(* Logix 5000 project; controller PLC_MCC1300_75F1 vendor 1 type 14 code 166 rev 32.11; software revision 32.04; part 49 of 83 *)
(* tags used below, declared in another part *)
   GP_ConversionXY : GP_ConversionXY;
   M30xTrimWheel : MAC_TrimmingWheels[5];
   M30xTrimWheel_HMR : MAC_TrimmingWheels_HMR[5];
   M30xTrimWheel_HMW : MAC_TrimmingWheels_HMW[5];
   M310B : MAC_Conveyor;
   M310B_ALM : MAC_Conveyor_ALM;
   M310B_Data : UDT_Convoy_SL;
   M310B_SpaceConv_Utilities : SpaceConv_Utilities;
   TMP_dIndex : DINT;
   TMP_rActualValue_cmm : REAL;
   xAlwaysON : BOOL;
   xDebugOFF : BOOL;
   Z401 : MAC_Zone;
(* MainProgram, continued *)

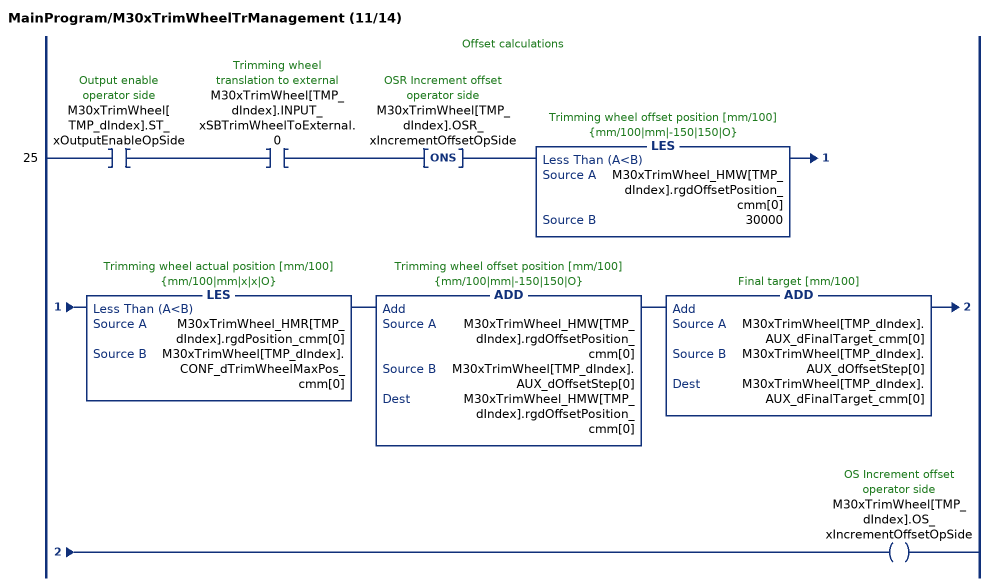
   [picture p745: MainProgram/M30xTrimWheelTrManagement rungs 25-25]
   // Offset calculations
   25: XIC(M30xTrimWheel[TMP_dIndex].ST_xOutputEnableOpSide)XIC(M30xTrimWheel[TMP_dIndex].INPUT_xSBTrimWheelToExternal.0)ONS(M30xTrimWheel[TMP_dIndex].OSR_xIncrementOffsetOpSide)LES(M30xTrimWheel_HMW[TMP_dIndex].rgdOffsetPosition_cmm[0],30000)LES(M30xTrimWheel_HMR[TMP_dIndex].rgdPosition_cmm[0],M30xTrimWheel[TMP_dIndex].CONF_dTrimWheelMaxPos_cmm[0])ADD(M30xTrimWheel_HMW[TMP_dIndex].rgdOffsetPosition_cmm[0],M30xTrimWheel[TMP_dIndex].AUX_dOffsetStep[0],M30xTrimWheel_HMW[TMP_dIndex].rgdOffsetPosition_cmm[0])ADD(M30xTrimWheel[TMP_dIndex].AUX_dFinalTarget_cmm[0],M30xTrimWheel[TMP_dIndex].AUX_dOffsetStep[0],M30xTrimWheel[TMP_dIndex].AUX_dFinalTarget_cmm[0])OTE(M30xTrimWheel[TMP_dIndex].OS_xIncrementOffsetOpSide);
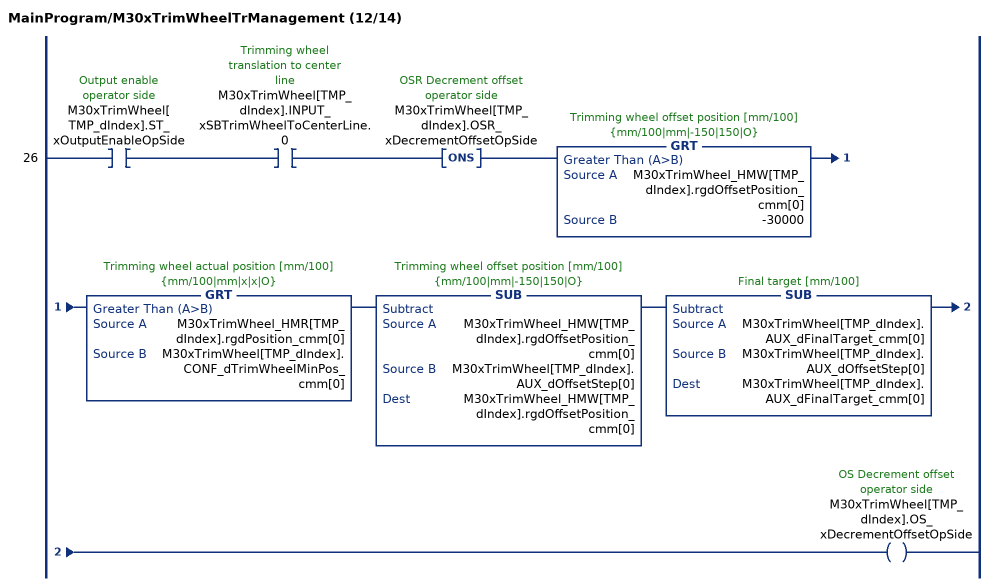
   26: XIC(M30xTrimWheel[TMP_dIndex].ST_xOutputEnableOpSide)XIC(M30xTrimWheel[TMP_dIndex].INPUT_xSBTrimWheelToCenterLine.0)ONS(M30xTrimWheel[TMP_dIndex].OSR_xDecrementOffsetOpSide)GRT(M30xTrimWheel_HMW[TMP_dIndex].rgdOffsetPosition_cmm[0],-30000)GRT(M30xTrimWheel_HMR[TMP_dIndex].rgdPosition_cmm[0],M30xTrimWheel[TMP_dIndex].CONF_dTrimWheelMinPos_cmm[0])SUB(M30xTrimWheel_HMW[TMP_dIndex].rgdOffsetPosition_cmm[0],M30xTrimWheel[TMP_dIndex].AUX_dOffsetStep[0],M30xTrimWheel_HMW[TMP_dIndex].rgdOffsetPosition_cmm[0])SUB(M30xTrimWheel[TMP_dIndex].AUX_dFinalTarget_cmm[0],M30xTrimWheel[TMP_dIndex].AUX_dOffsetStep[0],M30xTrimWheel[TMP_dIndex].AUX_dFinalTarget_cmm[0])OTE(M30xTrimWheel[TMP_dIndex].OS_xDecrementOffsetOpSide);
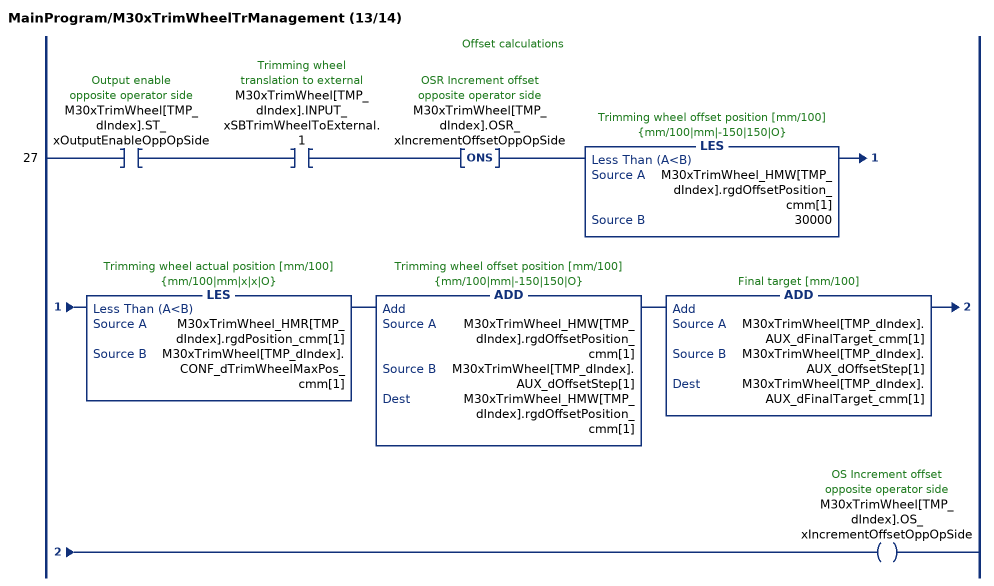
   // Offset calculations
   27: XIC(M30xTrimWheel[TMP_dIndex].ST_xOutputEnableOppOpSide)XIC(M30xTrimWheel[TMP_dIndex].INPUT_xSBTrimWheelToExternal.1)ONS(M30xTrimWheel[TMP_dIndex].OSR_xIncrementOffsetOppOpSide)LES(M30xTrimWheel_HMW[TMP_dIndex].rgdOffsetPosition_cmm[1],30000)LES(M30xTrimWheel_HMR[TMP_dIndex].rgdPosition_cmm[1],M30xTrimWheel[TMP_dIndex].CONF_dTrimWheelMaxPos_cmm[1])ADD(M30xTrimWheel_HMW[TMP_dIndex].rgdOffsetPosition_cmm[1],M30xTrimWheel[TMP_dIndex].AUX_dOffsetStep[1],M30xTrimWheel_HMW[TMP_dIndex].rgdOffsetPosition_cmm[1])ADD(M30xTrimWheel[TMP_dIndex].AUX_dFinalTarget_cmm[1],M30xTrimWheel[TMP_dIndex].AUX_dOffsetStep[1],M30xTrimWheel[TMP_dIndex].AUX_dFinalTarget_cmm[1])OTE(M30xTrimWheel[TMP_dIndex].OS_xIncrementOffsetOppOpSide);
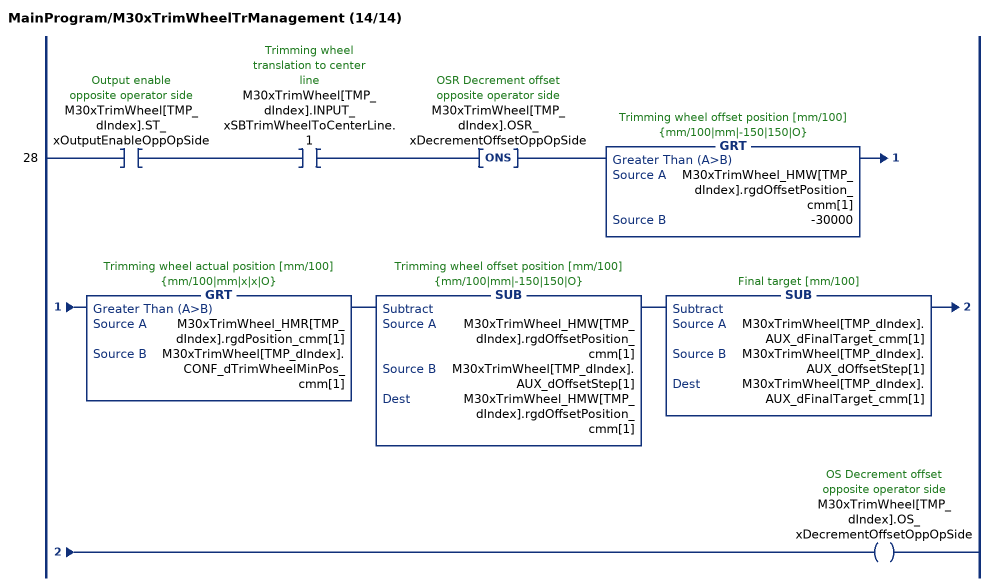
   28: XIC(M30xTrimWheel[TMP_dIndex].ST_xOutputEnableOppOpSide)XIC(M30xTrimWheel[TMP_dIndex].INPUT_xSBTrimWheelToCenterLine.1)ONS(M30xTrimWheel[TMP_dIndex].OSR_xDecrementOffsetOppOpSide)GRT(M30xTrimWheel_HMW[TMP_dIndex].rgdOffsetPosition_cmm[1],-30000)GRT(M30xTrimWheel_HMR[TMP_dIndex].rgdPosition_cmm[1],M30xTrimWheel[TMP_dIndex].CONF_dTrimWheelMinPos_cmm[1])SUB(M30xTrimWheel_HMW[TMP_dIndex].rgdOffsetPosition_cmm[1],M30xTrimWheel[TMP_dIndex].AUX_dOffsetStep[1],M30xTrimWheel_HMW[TMP_dIndex].rgdOffsetPosition_cmm[1])SUB(M30xTrimWheel[TMP_dIndex].AUX_dFinalTarget_cmm[1],M30xTrimWheel[TMP_dIndex].AUX_dOffsetStep[1],M30xTrimWheel[TMP_dIndex].AUX_dFinalTarget_cmm[1])OTE(M30xTrimWheel[TMP_dIndex].OS_xDecrementOffsetOppOpSide);
END_ROUTINE

ROUTINE M30xTrimWheelTrOppOpSide_Logic   (* ladder *)
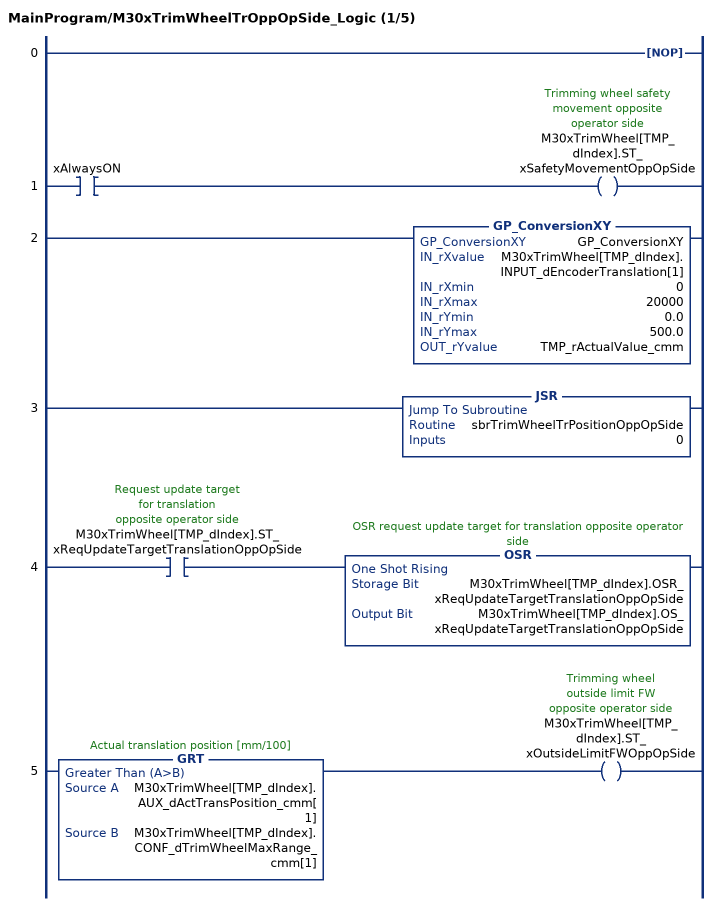
   0: NOP();
   1: XIC(xAlwaysON)OTE(M30xTrimWheel[TMP_dIndex].ST_xSafetyMovementOppOpSide);
   2: GP_ConversionXY(GP_ConversionXY,M30xTrimWheel[TMP_dIndex].INPUT_dEncoderTranslation[1],0,20000,0.0,500.0,TMP_rActualValue_cmm);
   3: JSR(sbrTrimWheelTrPositionOppOpSide,0);
   4: XIC(M30xTrimWheel[TMP_dIndex].ST_xReqUpdateTargetTranslationOppOpSide)OSR(M30xTrimWheel[TMP_dIndex].OSR_xReqUpdateTargetTranslationOppOpSide,M30xTrimWheel[TMP_dIndex].OS_xReqUpdateTargetTranslationOppOpSide);
   5: GRT(M30xTrimWheel[TMP_dIndex].AUX_dActTransPosition_cmm[1],M30xTrimWheel[TMP_dIndex].CONF_dTrimWheelMaxRange_cmm[1])OTE(M30xTrimWheel[TMP_dIndex].ST_xOutsideLimitFWOppOpSide);
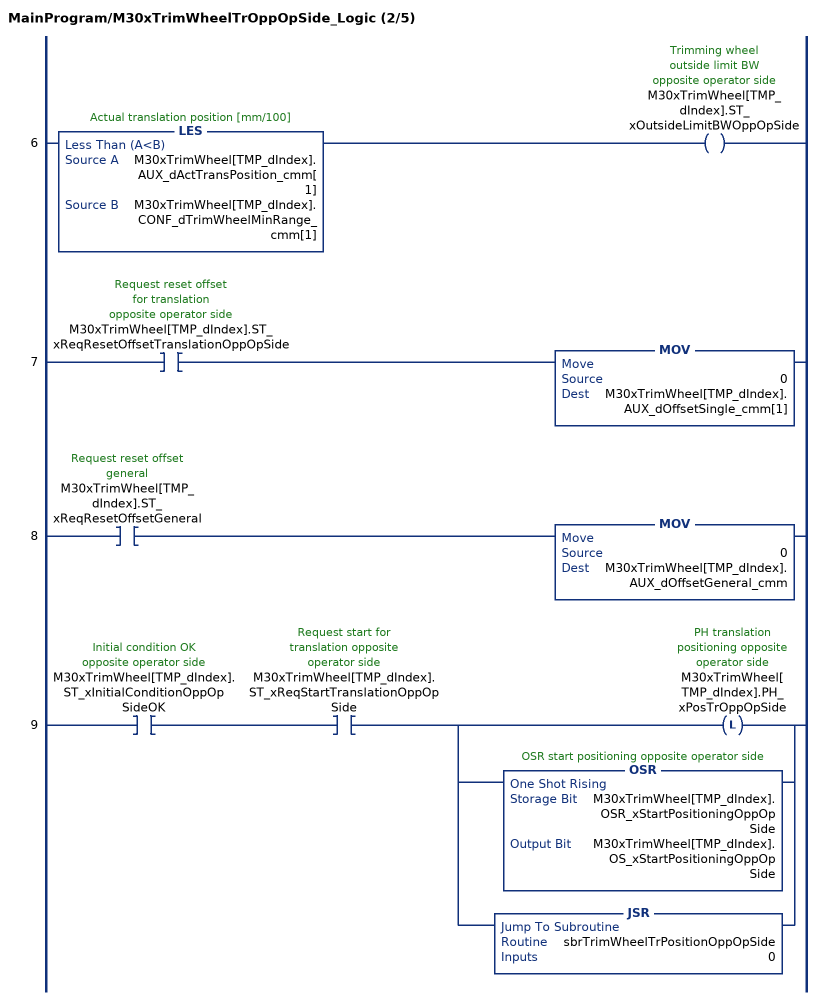
   6: LES(M30xTrimWheel[TMP_dIndex].AUX_dActTransPosition_cmm[1],M30xTrimWheel[TMP_dIndex].CONF_dTrimWheelMinRange_cmm[1])OTE(M30xTrimWheel[TMP_dIndex].ST_xOutsideLimitBWOppOpSide);
   7: XIC(M30xTrimWheel[TMP_dIndex].ST_xReqResetOffsetTranslationOppOpSide)MOV(0,M30xTrimWheel[TMP_dIndex].AUX_dOffsetSingle_cmm[1]);
   8: XIC(M30xTrimWheel[TMP_dIndex].ST_xReqResetOffsetGeneral)MOV(0,M30xTrimWheel[TMP_dIndex].AUX_dOffsetGeneral_cmm);
   9: XIC(M30xTrimWheel[TMP_dIndex].ST_xInitialConditionOppOpSideOK)XIC(M30xTrimWheel[TMP_dIndex].ST_xReqStartTranslationOppOpSide)[OTL(M30xTrimWheel[TMP_dIndex].PH_xPosTrOppOpSide) ,OSR(M30xTrimWheel[TMP_dIndex].OSR_xStartPositioningOppOpSide,M30xTrimWheel[TMP_dIndex].OS_xStartPositioningOppOpSide) ,JSR(sbrTrimWheelTrPositionOppOpSide,0) ];
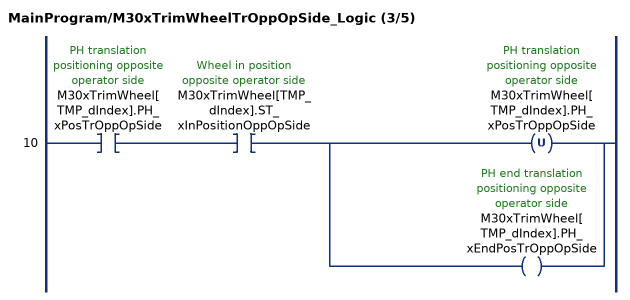
   10: XIC(M30xTrimWheel[TMP_dIndex].PH_xPosTrOppOpSide)XIC(M30xTrimWheel[TMP_dIndex].ST_xInPositionOppOpSide)[OTU(M30xTrimWheel[TMP_dIndex].PH_xPosTrOppOpSide) ,OTE(M30xTrimWheel[TMP_dIndex].PH_xEndPosTrOppOpSide) ];
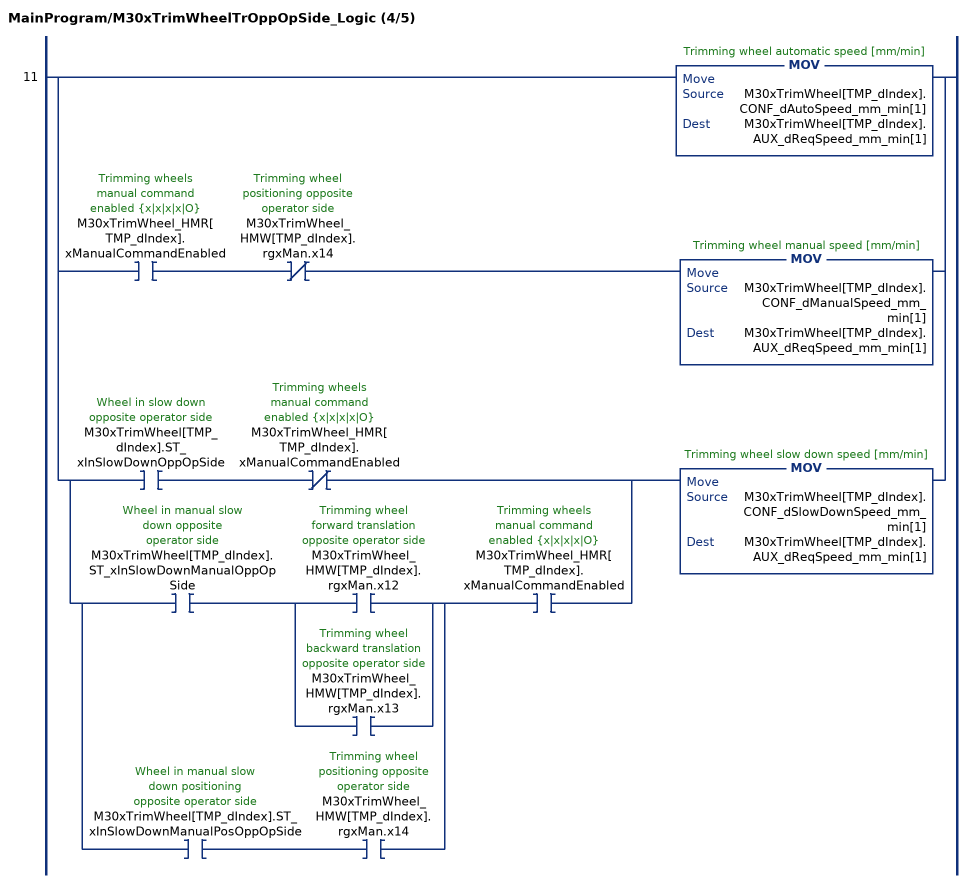
   11: [MOV(M30xTrimWheel[TMP_dIndex].CONF_dAutoSpeed_mm_min[1],M30xTrimWheel[TMP_dIndex].AUX_dReqSpeed_mm_min[1]) ,XIC(M30xTrimWheel_HMR[TMP_dIndex].xManualCommandEnabled) XIO(M30xTrimWheel_HMW[TMP_dIndex].rgxMan.x14) MOV(M30xTrimWheel[TMP_dIndex].CONF_dManualSpeed_mm_min[1],M30xTrimWheel[TMP_dIndex].AUX_dReqSpeed_mm_min[1]) ,[XIC(M30xTrimWheel[TMP_dIndex].ST_xInSlowDownOppOpSide) XIO(M30xTrimWheel_HMR[TMP_dIndex].xManualCommandEnabled) ,[XIC(M30xTrimWheel[TMP_dIndex].ST_xInSlowDownManualOppOpSide) [XIC(M30xTrimWheel_HMW[TMP_dIndex].rgxMan.x12) ,XIC(M30xTrimWheel_HMW[TMP_dIndex].rgxMan.x13) ] ,XIC(M30xTrimWheel[TMP_dIndex].ST_xInSlowDownManualPosOppOpSide) XIC(M30xTrimWheel_HMW[TMP_dIndex].rgxMan.x14) ] XIC(M30xTrimWheel_HMR[TMP_dIndex].xManualCommandEnabled) ] MOV(M30xTrimWheel[TMP_dIndex].CONF_dSlowDownSpeed_mm_min[1],M30xTrimWheel[TMP_dIndex].AUX_dReqSpeed_mm_min[1]) ];
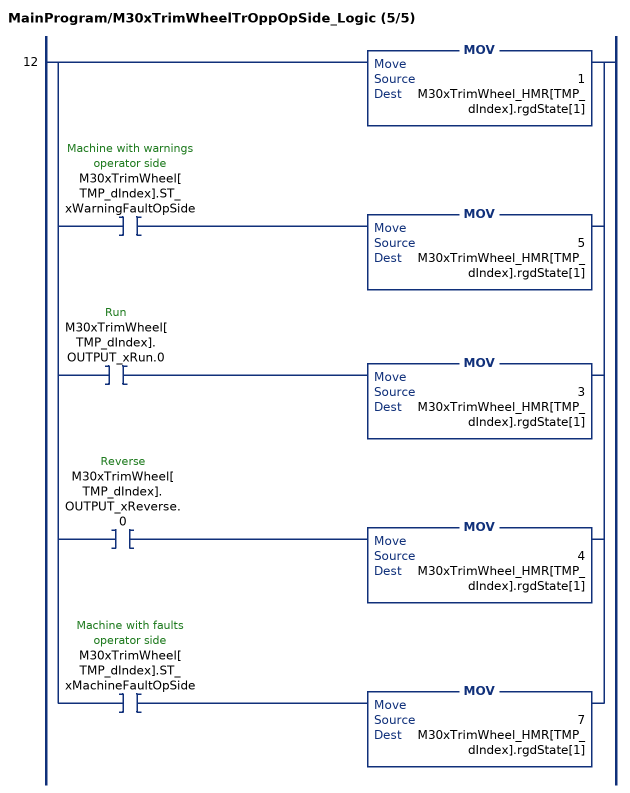
   12: [MOV(1,M30xTrimWheel_HMR[TMP_dIndex].rgdState[1]) ,XIC(M30xTrimWheel[TMP_dIndex].ST_xWarningFaultOpSide) MOV(5,M30xTrimWheel_HMR[TMP_dIndex].rgdState[1]) ,XIC(M30xTrimWheel[TMP_dIndex].OUTPUT_xRun.0) MOV(3,M30xTrimWheel_HMR[TMP_dIndex].rgdState[1]) ,XIC(M30xTrimWheel[TMP_dIndex].OUTPUT_xReverse.0) MOV(4,M30xTrimWheel_HMR[TMP_dIndex].rgdState[1]) ,XIC(M30xTrimWheel[TMP_dIndex].ST_xMachineFaultOpSide) MOV(7,M30xTrimWheel_HMR[TMP_dIndex].rgdState[1]) ];
END_ROUTINE

ROUTINE M30xTrimWheelTrOpSide_Logic   (* ladder *)
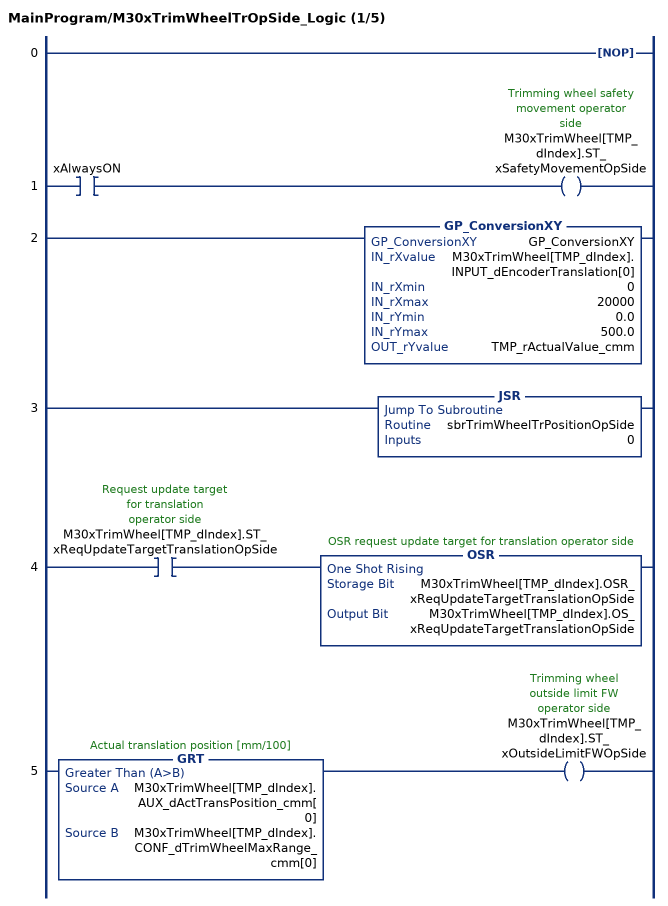
   0: NOP();
   1: XIC(xAlwaysON)OTE(M30xTrimWheel[TMP_dIndex].ST_xSafetyMovementOpSide);
   2: GP_ConversionXY(GP_ConversionXY,M30xTrimWheel[TMP_dIndex].INPUT_dEncoderTranslation[0],0,20000,0.0,500.0,TMP_rActualValue_cmm);
   3: JSR(sbrTrimWheelTrPositionOpSide,0);
   4: XIC(M30xTrimWheel[TMP_dIndex].ST_xReqUpdateTargetTranslationOpSide)OSR(M30xTrimWheel[TMP_dIndex].OSR_xReqUpdateTargetTranslationOpSide,M30xTrimWheel[TMP_dIndex].OS_xReqUpdateTargetTranslationOpSide);
   5: GRT(M30xTrimWheel[TMP_dIndex].AUX_dActTransPosition_cmm[0],M30xTrimWheel[TMP_dIndex].CONF_dTrimWheelMaxRange_cmm[0])OTE(M30xTrimWheel[TMP_dIndex].ST_xOutsideLimitFWOpSide);
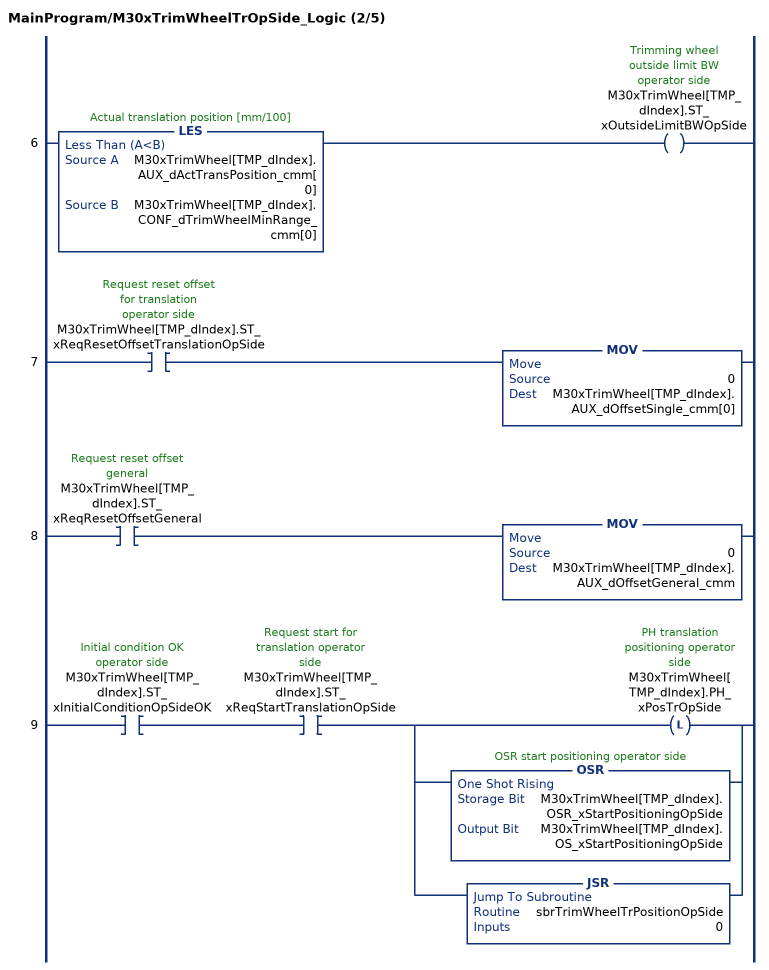
   6: LES(M30xTrimWheel[TMP_dIndex].AUX_dActTransPosition_cmm[0],M30xTrimWheel[TMP_dIndex].CONF_dTrimWheelMinRange_cmm[0])OTE(M30xTrimWheel[TMP_dIndex].ST_xOutsideLimitBWOpSide);
   7: XIC(M30xTrimWheel[TMP_dIndex].ST_xReqResetOffsetTranslationOpSide)MOV(0,M30xTrimWheel[TMP_dIndex].AUX_dOffsetSingle_cmm[0]);
   8: XIC(M30xTrimWheel[TMP_dIndex].ST_xReqResetOffsetGeneral)MOV(0,M30xTrimWheel[TMP_dIndex].AUX_dOffsetGeneral_cmm);
   9: XIC(M30xTrimWheel[TMP_dIndex].ST_xInitialConditionOpSideOK)XIC(M30xTrimWheel[TMP_dIndex].ST_xReqStartTranslationOpSide)[OTL(M30xTrimWheel[TMP_dIndex].PH_xPosTrOpSide) ,OSR(M30xTrimWheel[TMP_dIndex].OSR_xStartPositioningOpSide,M30xTrimWheel[TMP_dIndex].OS_xStartPositioningOpSide) ,JSR(sbrTrimWheelTrPositionOpSide,0) ];
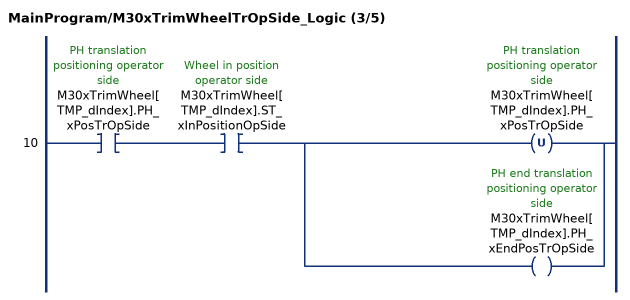
   10: XIC(M30xTrimWheel[TMP_dIndex].PH_xPosTrOpSide)XIC(M30xTrimWheel[TMP_dIndex].ST_xInPositionOpSide)[OTU(M30xTrimWheel[TMP_dIndex].PH_xPosTrOpSide) ,OTE(M30xTrimWheel[TMP_dIndex].PH_xEndPosTrOpSide) ];
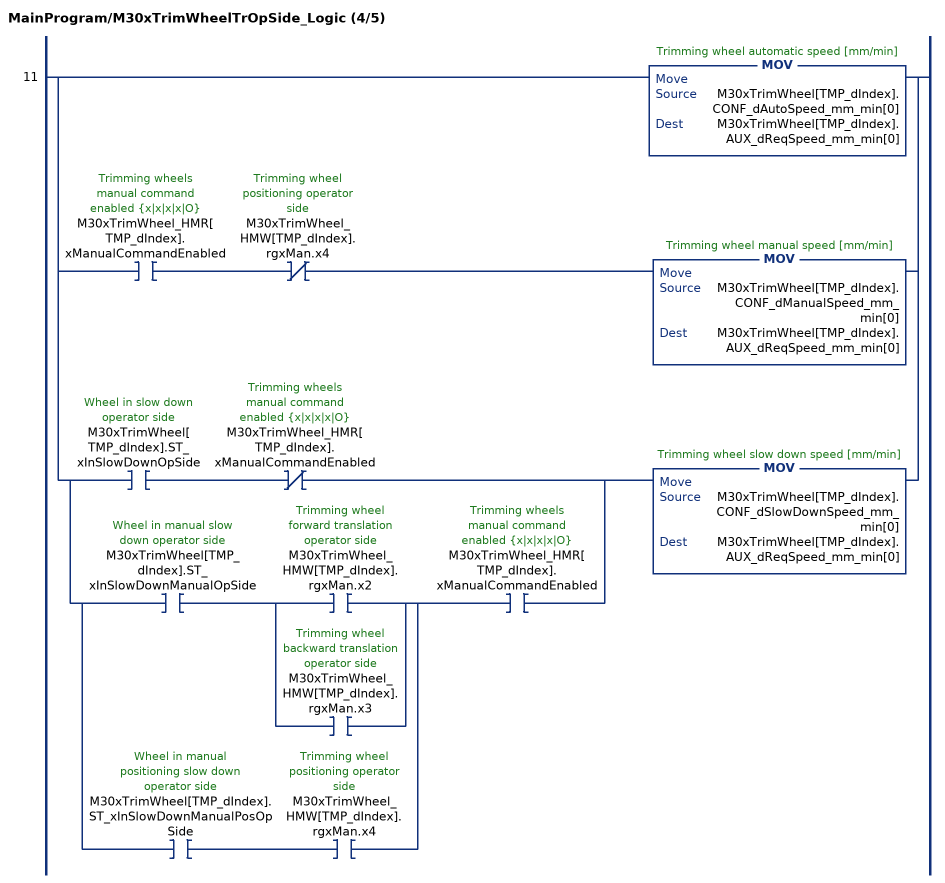
   11: [MOV(M30xTrimWheel[TMP_dIndex].CONF_dAutoSpeed_mm_min[0],M30xTrimWheel[TMP_dIndex].AUX_dReqSpeed_mm_min[0]) ,XIC(M30xTrimWheel_HMR[TMP_dIndex].xManualCommandEnabled) XIO(M30xTrimWheel_HMW[TMP_dIndex].rgxMan.x4) MOV(M30xTrimWheel[TMP_dIndex].CONF_dManualSpeed_mm_min[0],M30xTrimWheel[TMP_dIndex].AUX_dReqSpeed_mm_min[0]) ,[XIC(M30xTrimWheel[TMP_dIndex].ST_xInSlowDownOpSide) XIO(M30xTrimWheel_HMR[TMP_dIndex].xManualCommandEnabled) ,[XIC(M30xTrimWheel[TMP_dIndex].ST_xInSlowDownManualOpSide) [XIC(M30xTrimWheel_HMW[TMP_dIndex].rgxMan.x2) ,XIC(M30xTrimWheel_HMW[TMP_dIndex].rgxMan.x3) ] ,XIC(M30xTrimWheel[TMP_dIndex].ST_xInSlowDownManualPosOpSide) XIC(M30xTrimWheel_HMW[TMP_dIndex].rgxMan.x4) ] XIC(M30xTrimWheel_HMR[TMP_dIndex].xManualCommandEnabled) ] MOV(M30xTrimWheel[TMP_dIndex].CONF_dSlowDownSpeed_mm_min[0],M30xTrimWheel[TMP_dIndex].AUX_dReqSpeed_mm_min[0]) ];
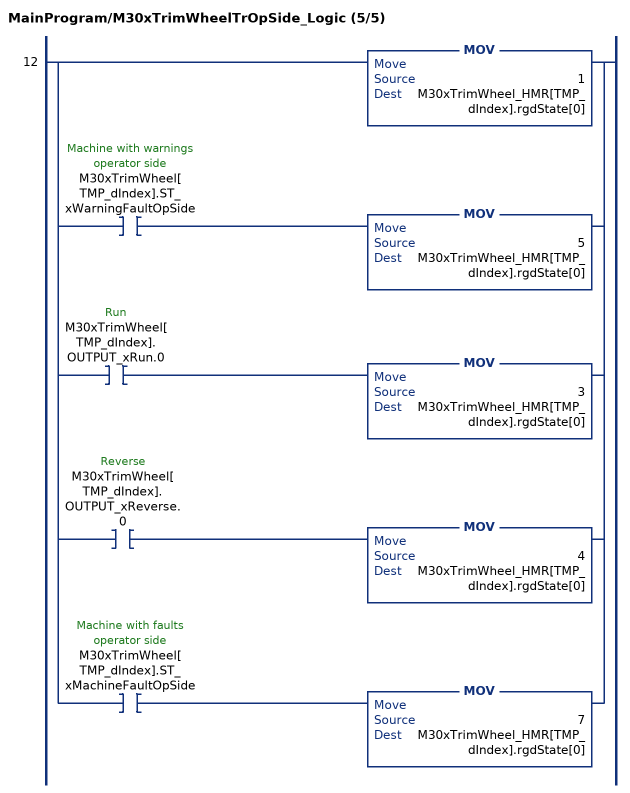
   12: [MOV(1,M30xTrimWheel_HMR[TMP_dIndex].rgdState[0]) ,XIC(M30xTrimWheel[TMP_dIndex].ST_xWarningFaultOpSide) MOV(5,M30xTrimWheel_HMR[TMP_dIndex].rgdState[0]) ,XIC(M30xTrimWheel[TMP_dIndex].OUTPUT_xRun.0) MOV(3,M30xTrimWheel_HMR[TMP_dIndex].rgdState[0]) ,XIC(M30xTrimWheel[TMP_dIndex].OUTPUT_xReverse.0) MOV(4,M30xTrimWheel_HMR[TMP_dIndex].rgdState[0]) ,XIC(M30xTrimWheel[TMP_dIndex].ST_xMachineFaultOpSide) MOV(7,M30xTrimWheel_HMR[TMP_dIndex].rgdState[0]) ];
END_ROUTINE

ROUTINE M310B_Alarm   (* ladder *)
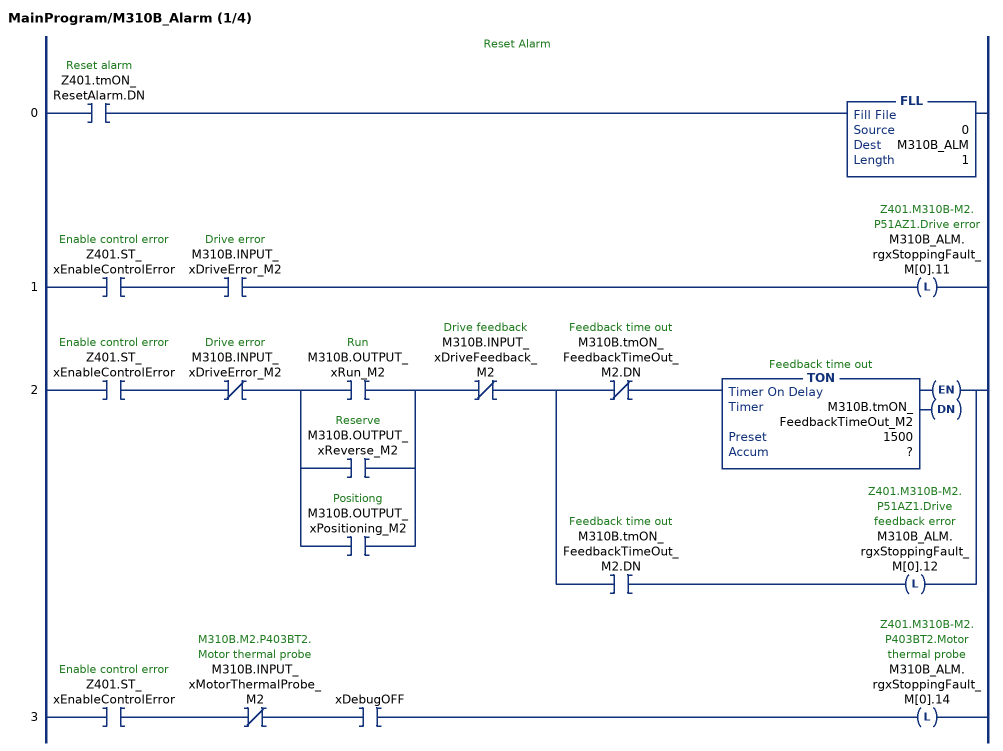
   // Reset Alarm
   0: XIC(Z401.tmON_ResetAlarm.DN)FLL(0,M310B_ALM,1);
   1: XIC(Z401.ST_xEnableControlError)XIC(M310B.INPUT_xDriveError_M2)OTL(M310B_ALM.rgxStoppingFault_M[0].11);
   2: XIC(Z401.ST_xEnableControlError)XIO(M310B.INPUT_xDriveError_M2)[XIC(M310B.OUTPUT_xRun_M2) ,XIC(M310B.OUTPUT_xReverse_M2) ,XIC(M310B.OUTPUT_xPositioning_M2) ]XIO(M310B.INPUT_xDriveFeedback_M2)[XIO(M310B.tmON_FeedbackTimeOut_M2.DN) TON(M310B.tmON_FeedbackTimeOut_M2,?,?) ,XIC(M310B.tmON_FeedbackTimeOut_M2.DN) OTL(M310B_ALM.rgxStoppingFault_M[0].12) ];
   3: XIC(Z401.ST_xEnableControlError)XIO(M310B.INPUT_xMotorThermalProbe_M2)XIC(xDebugOFF)OTL(M310B_ALM.rgxStoppingFault_M[0].14);
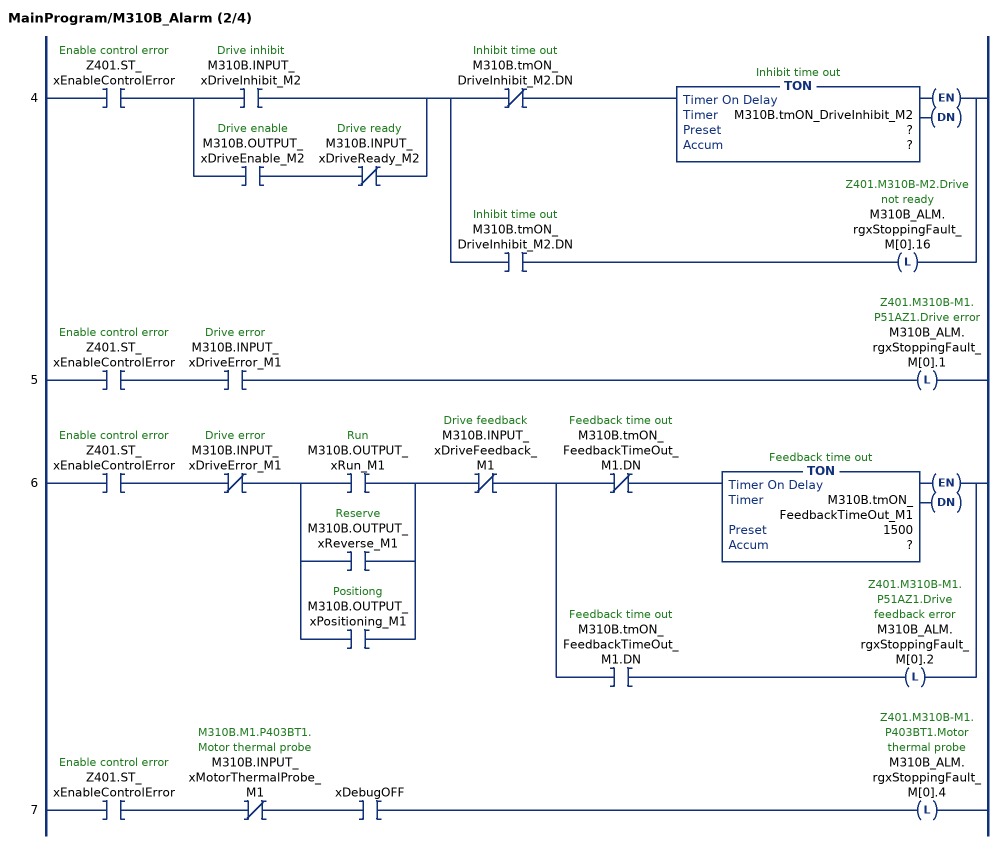
   4: XIC(Z401.ST_xEnableControlError)[XIC(M310B.INPUT_xDriveInhibit_M2) ,XIC(M310B.OUTPUT_xDriveEnable_M2) XIO(M310B.INPUT_xDriveReady_M2) ][XIO(M310B.tmON_DriveInhibit_M2.DN) TON(M310B.tmON_DriveInhibit_M2,?,?) ,XIC(M310B.tmON_DriveInhibit_M2.DN) OTL(M310B_ALM.rgxStoppingFault_M[0].16) ];
   5: XIC(Z401.ST_xEnableControlError)XIC(M310B.INPUT_xDriveError_M1)OTL(M310B_ALM.rgxStoppingFault_M[0].1);
   6: XIC(Z401.ST_xEnableControlError)XIO(M310B.INPUT_xDriveError_M1)[XIC(M310B.OUTPUT_xRun_M1) ,XIC(M310B.OUTPUT_xReverse_M1) ,XIC(M310B.OUTPUT_xPositioning_M1) ]XIO(M310B.INPUT_xDriveFeedback_M1)[XIO(M310B.tmON_FeedbackTimeOut_M1.DN) TON(M310B.tmON_FeedbackTimeOut_M1,?,?) ,XIC(M310B.tmON_FeedbackTimeOut_M1.DN) OTL(M310B_ALM.rgxStoppingFault_M[0].2) ];
   7: XIC(Z401.ST_xEnableControlError)XIO(M310B.INPUT_xMotorThermalProbe_M1)XIC(xDebugOFF)OTL(M310B_ALM.rgxStoppingFault_M[0].4);
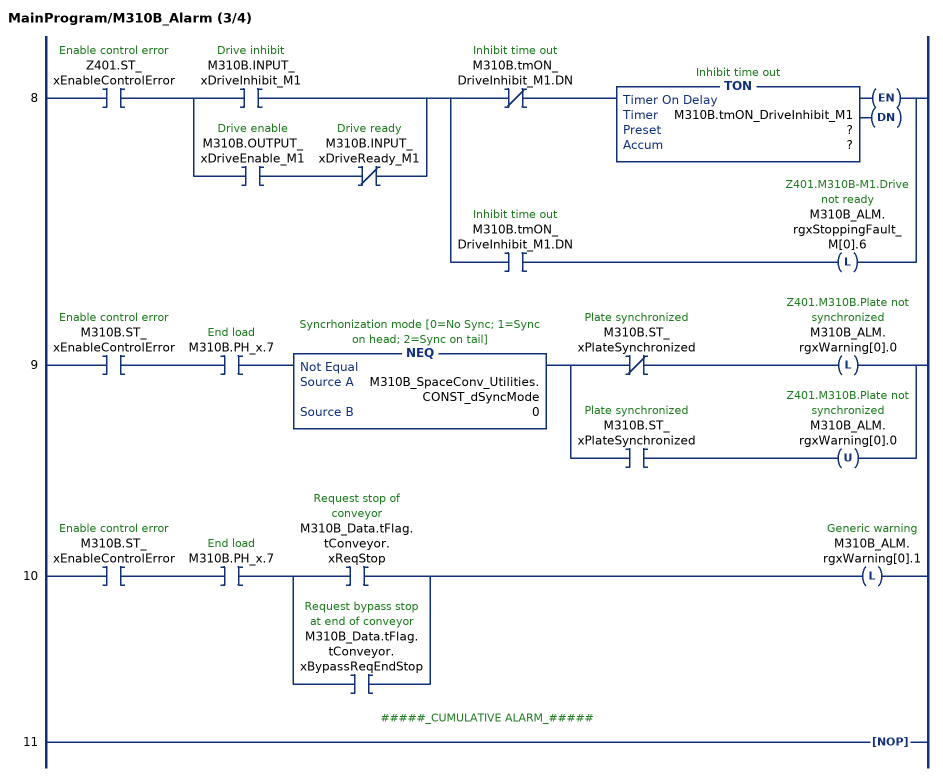
   8: XIC(Z401.ST_xEnableControlError)[XIC(M310B.INPUT_xDriveInhibit_M1) ,XIC(M310B.OUTPUT_xDriveEnable_M1) XIO(M310B.INPUT_xDriveReady_M1) ][XIO(M310B.tmON_DriveInhibit_M1.DN) TON(M310B.tmON_DriveInhibit_M1,?,?) ,XIC(M310B.tmON_DriveInhibit_M1.DN) OTL(M310B_ALM.rgxStoppingFault_M[0].6) ];
   9: XIC(M310B.ST_xEnableControlError)XIC(M310B.PH_x.7)NEQ(M310B_SpaceConv_Utilities.CONST_dSyncMode,0)[XIO(M310B.ST_xPlateSynchronized) OTL(M310B_ALM.rgxWarning[0].0) ,XIC(M310B.ST_xPlateSynchronized) OTU(M310B_ALM.rgxWarning[0].0) ];
   10: XIC(M310B.ST_xEnableControlError)XIC(M310B.PH_x.7)[XIC(M310B_Data.tFlag.tConveyor.xReqStop) ,XIC(M310B_Data.tFlag.tConveyor.xBypassReqEndStop) ]OTL(M310B_ALM.rgxWarning[0].1);
   // #####_CUMULATIVE ALARM_#####
   11: NOP();
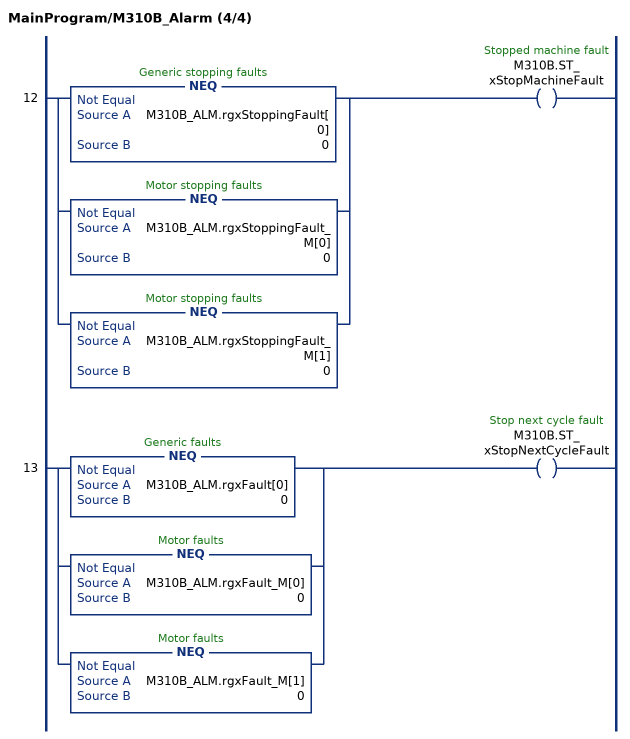
   12: [NEQ(M310B_ALM.rgxStoppingFault[0],0) ,NEQ(M310B_ALM.rgxStoppingFault_M[0],0) ,NEQ(M310B_ALM.rgxStoppingFault_M[1],0) ]OTE(M310B.ST_xStopMachineFault);
   13: [NEQ(M310B_ALM.rgxFault[0],0) ,NEQ(M310B_ALM.rgxFault_M[0],0) ,NEQ(M310B_ALM.rgxFault_M[1],0) ]OTE(M310B.ST_xStopNextCycleFault);
END_ROUTINE
